// TIA Portal project "PalletizerLine" (V17)

(* hardware
DEVICE "S7-1500 station"  S7-1500 station
   slot 0: "Rail_0"  Rack  6ES7 590-1***0-0AA0
   slot 0: "PM 70W 120/230VAC"  PM 70W 120/230VAC  6EP1332-4BA00
   slot 1: "PLC_1"  CPU 1511-1 PN  6ES7 511-1AK02-0AB0  V2.9
      slot 3: "CPU display_1"  6ES7591-1AA00-0AA0
      slot 32768: "PROFINET interface_1"  X1
      slot 34817: "Virtual CP interface port_1"  Virtual CP interface port  Virtual CP interface port
   slot 2: "AI 8xU/I/RTD/TC ST_1"  AI 8xU/I/RTD/TC ST  6ES7 531-7KF00-0AB0  V2.2
   slot 3: "AI 8xU/I/RTD/TC ST_2"  AI 8xU/I/RTD/TC ST  6ES7 531-7KF00-0AB0  V2.2
   slot 4: "AI 8xU/I/RTD/TC ST_3"  AI 8xU/I/RTD/TC ST  6ES7 531-7KF00-0AB0  V2.2
   slot 5: "AI 8xU/I/RTD/TC ST_4"  AI 8xU/I/RTD/TC ST  6ES7 531-7KF00-0AB0  V2.2
   slot 6: "DI 16x24VDC BA_1"  DI 16x24VDC BA  6ES7 521-1BH10-0AA0  V1.1
DEVICE "HMI_TP1200"  TP1200 Comfort
   slot 0: "TP1200 Comfort"  TP1200 Comfort  6AV2 124-0MC01-0AX0  14.0.1.0
   slot 1: "HMI_RT_1"  TP1200 Comfort  6AV2 124-0MC01-0AX0  14.0.1.0
   slot 5: "Labeler HMI_TP1200.HMI.1"  PROFINET Interface  IE_CP  14.0.1.0
      slot 1: "PROFINET_Interface_1"  PROFINET Interface
         slot 1: "PORT_1"  Port  1.0.0.0
         slot 2: "PORT_2"  Port  1.0.0.0
   slot 7: "Labeler HMI_TP1200.HMI._CP_1"  MPI/DP Interface  MPI-DP_CP  14.0.1.0
*)

// ===== PLC "PLC_1"  CPU 1511-1 PN =====

VAR_GLOBAL   // PLC tag table "Default tag table"
   "System_Byte" AT %MB0 : Byte;   // System byte
   "FirstScan" AT %M0.0 : Bool;   // First scan PLC
   "DiagStatusUpdate" AT %M0.1 : Bool;   // Diagnostic status PLC updated
   "AlwaysTRUE" AT %M0.2 : Bool;   // Bit always true
   "AlwaysFALSE" AT %M0.3 : Bool;   // Bit always false
   "Clock_Byte" AT %MB1 : Byte;   // Clock byte
   "Clock_10Hz" AT %M1.0 : Bool;   // Clock pulse period 0,1s
   "Clock_5Hz" AT %M1.1 : Bool;   // Clock pulse period 0,2s
   "Clock_2.5Hz" AT %M1.2 : Bool;   // Clock pulse period 0,4s
   "Clock_2Hz" AT %M1.3 : Bool;   // Clock pulse period 0,5s
   "Clock_1.25Hz" AT %M1.4 : Bool;   // Clock pulse period 0,8s
   "Clock_1Hz" AT %M1.5 : Bool;   // Clock pulse period 1s
   "Clock_0.625Hz" AT %M1.6 : Bool;   // Clock pulse period 1,6s
   "Clock_0.5Hz" AT %M1.7 : Bool;   // Clock pulse period 2s
   "Tag_1" AT %I0.0 : Bool;
   "Tag_2" AT %Q0.0 : Bool;
   "Tag_3" AT %I0.1 : Bool;
   "Tag_4" AT %Q0.1 : Bool;
   "Tag_5" AT %Q0.2 : Bool;
   "Tag_6" AT %Q0.3 : Bool;
   "Tag_7" AT %Q0.4 : Bool;
   "Tag_8" AT %I0.2 : Bool;
   "Tag_9" AT %Q0.5 : Bool;
   "Tag_10" AT %I0.3 : Bool;
   "Tag_11" AT %Q0.6 : Bool;
   "Tag_12" AT %I0.4 : Bool;
   "Tag_13" AT %I0.5 : Bool;
   "Tag_14" AT %I0.6 : Bool;
   "Tag_15" AT %I0.7 : Bool;
   "Tag_16" AT %I1.0 : Bool;
   "Tag_17" AT %I1.1 : Bool;
   "Tag_18" AT %I1.2 : Bool;
   "Tag_19" AT %Q0.7 : Bool;
   "Tag_20" AT %Q1.0 : Bool;
   "Tag_21" AT %Q1.1 : Bool;
   "Tag_22" AT %Q1.2 : Bool;
   "Tag_23" AT %Q1.3 : Bool;
   "Tag_24" AT %Q1.4 : Bool;
   "Tag_25" AT %Q1.5 : Bool;
   "Tag_26" AT %Q1.6 : Bool;
   "Tag_27" AT %Q1.7 : Bool;
   "Tag_28" AT %Q2.0 : Bool;
   "Tag_29" AT %Q2.1 : Bool;
   "Tag_30" AT %Q2.2 : Bool;
   "Tag_31" AT %Q2.3 : Bool;
END_VAR

VAR_GLOBAL CONSTANT   // PLC tag table "CPG_Constants"
   "CPG_NO_OF_ELEMENTS_EVENT_STATUS_UPPER_LIM" : Int := 29;   // Number of Alarms, Warning and PackML Status events used by Event Status UDT (Array size of 0..x)
   "CPG_NO_OF_ADMIN_EVENTS_UPPER_LIM" : Int := 9;   // Number of Alarms and Warning events found in the PackTags Admin Area - active alarms / warnings. (Array size of 0..x)
   "CPG_NO_OF_ADMIN_EVENTS_HISTORY_UPPER_LIM" : Int := 9;   // Number of Alarms and Warning events found in the PackTags Admin Area - historical alarms / warnings. (Array size of 0..x)
   "CPG_NO_OF_PROD_CONSUMED_COUNT_UPPER_LIM" : Int := 0;   // Number of Prod Consumed Counter Array Size (PackTags Admin) (Array size of 0..x)
   "CPG_NO_OF_PROD_PROCESSED_COUNT_UPPER_LIM" : Int := 0;   // Number of Prod Processed Counter Array Size (PackTags Admin) (Array size of 0..x)
   "CPG_NO_OF_PROD_DEFECTIVE_COUNT_UPPER_LIM" : Int := 0;   // Number of Prod Defective Counter Array Size (PackTags Admin) (Array size of 0..x)
   "CPG_NO_OF_STS_ELEMENTS_EVENT_SUM_UPPER_LIM" : Int := 99;   // Number of Alarms, Warning and PackML Status events used by Event Summation UDT (Array size of 0..x)
   "CPG_NO_OF_HMI_SORT_EVENTS_UPPER_LIM" : Int := 19;   // Number of Alarms and Warning events found for the HMI area - sorted HMI alarms / warnings. (Array size of 0..x)
   "CPG_NO_OF_CFG_ALARMS_UPPER_LIM" : Int := 39;   // Number of Cfg Alarm event configurations (Array size of 0..x)
   "CPG_NO_OF_CFG_WARNINGS_UPPER_LIM" : Int := 29;   // Number of Cfg Warning event configurations (Array size of 0..x)
   "CPG_NO_OF_CFG_STATUS_UPPER_LIM" : Int := 19;   // Number of Cfg Status event configurations (Array size of 0..x)
   "CPG_NO_OF_STATUS_PARAMETERS_UPPER_LIM" : Int := 0;   // Number of Status Parameters (Array size of 0..x)
   "CPG_NO_OF_COMMAND_PARAMETERS_UPPER_LIM" : Int := 0;   // Number of Command Parameters (Array size of 0..x)
   "CPG_NO_OF_ADMIN_PARAMETERS_UPPER_LIM" : Int := 0;   // Number of Admin Parameters (Array size of 0..x)
   "CPG_NO_OF_RECIPE_UPPER_LIM" : Int := 20;   // Number of Project Recipies (Array size of 0..x)
   "CPG_NO_OF_SETPOINT_REAL_UPPER_LIM" : Int := 0;   // Number of Setpoints with a REAL type (Array size of 0..x)
   "CPG_NO_OF_SETPOINT_DINT_UPPER_LIM" : Int := 0;   // Number of Setpoints with a DINT type (Array size of 0..x)
   "CPG_NO_OF_SETPOINT_BOOL_UPPER_LIM" : Int := 0;   // Number of Setpoints with a BOOL type (Array size of 0..x)
   "CPG_NO_OF_SETPOINT_STRING_UPPER_LIM" : Int := 0;   // Number of Setpoints with a STRING type (Array size of 0..x)
   "CPG_PARTEO_NO_OF_ERRORS_UPPER_LIM" : Int := 100;   // Number of Unique Error IDs tracked by PARETO Error Blocks
END_VAR

VAR_GLOBAL CONSTANT   // PLC tag table "LPMLV30_Constants"
   "LPMLV30_MODE_INVALID" : DInt := 0;   // OMAC PackMLV30 unit mode Invalid
   "LPMLV30_MODE_PRODUCTION" : DInt := 1;   // OMAC PackMLV30 unit mode Production
   "LPMLV30_MODE_MAINTENANCE" : DInt := 2;   // OMAC PackMLV30 unit mode Maintenance
   "LPMLV30_MODE_MANUAL" : DInt := 3;   // OMAC PackMLV30 unit mode Manual
   "LPMLV30_MODE_USER_01" : DInt := 4;   // OMAC PackMLV30 user-defined unit mode 01
   "LPMLV30_MODE_USER_02" : DInt := 5;   // OMAC PackMLV30 user-defined unit mode 02
   "LPMLV30_MODE_USER_03" : DInt := 6;   // OMAC PackMLV30 user-defined unit mode 03
   "LPMLV30_MODE_USER_04" : DInt := 7;   // OMAC PackMLV30 user-defined unit mode 04
   "LPMLV30_MODE_USER_05" : DInt := 8;   // OMAC PackMLV30 user-defined unit mode 05
   "LPMLV30_MODE_USER_06" : DInt := 9;   // OMAC PackMLV30 user-defined unit mode 06
   "LPMLV30_MODE_USER_07" : DInt := 10;   // OMAC PackMLV30 user-defined unit mode 07
   "LPMLV30_MODE_USER_08" : DInt := 11;   // OMAC PackMLV30 user-defined unit mode 08
   "LPMLV30_MODE_USER_09" : DInt := 12;   // OMAC PackMLV30 user-defined unit mode 09
   "LPMLV30_MODE_USER_10" : DInt := 13;   // OMAC PackMLV30 user-defined unit mode 10
   "LPMLV30_MODE_USER_11" : DInt := 14;   // OMAC PackMLV30 user-defined unit mode 11
   "LPMLV30_MODE_USER_12" : DInt := 15;   // OMAC PackMLV30 user-defined unit mode 12
   "LPMLV30_MODE_USER_13" : DInt := 16;   // OMAC PackMLV30 user-defined unit mode 13
   "LPMLV30_MODE_USER_14" : DInt := 17;   // OMAC PackMLV30 user-defined unit mode 14
   "LPMLV30_MODE_USER_15" : DInt := 18;   // OMAC PackMLV30 user-defined unit mode 15
   "LPMLV30_MODE_USER_16" : DInt := 19;   // OMAC PackMLV30 user-defined unit mode 16
   "LPMLV30_MODE_USER_17" : DInt := 20;   // OMAC PackMLV30 user-defined unit mode 17
   "LPMLV30_MODE_USER_18" : DInt := 21;   // OMAC PackMLV30 user-defined unit mode 18
   "LPMLV30_MODE_USER_19" : DInt := 22;   // OMAC PackMLV30 user-defined unit mode 19
   "LPMLV30_MODE_USER_20" : DInt := 23;   // OMAC PackMLV30 user-defined unit mode 20
   "LPMLV30_MODE_USER_21" : DInt := 24;   // OMAC PackMLV30 user-defined unit mode 21
   "LPMLV30_MODE_USER_22" : DInt := 25;   // OMAC PackMLV30 user-defined unit mode 22
   "LPMLV30_MODE_USER_23" : DInt := 26;   // OMAC PackMLV30 user-defined unit mode 23
   "LPMLV30_MODE_USER_24" : DInt := 27;   // OMAC PackMLV30 user-defined unit mode 24
   "LPMLV30_MODE_USER_25" : DInt := 28;   // OMAC PackMLV30 user-defined unit mode 25
   "LPMLV30_MODE_USER_26" : DInt := 29;   // OMAC PackMLV30 user-defined unit mode 26
   "LPMLV30_MODE_USER_27" : DInt := 30;   // OMAC PackMLV30 user-defined unit mode 27
   "LPMLV30_MODE_USER_28" : DInt := 31;   // OMAC PackMLV30 user-defined unit mode 28
   "LPMLV30_STATE_UNDEFINED" : DInt := 0;   // OMAC PackMLV30 state Undefined
   "LPMLV30_STATE_CLEARING" : DInt := 1;   // OMAC PackMLV30 state Clearing
   "LPMLV30_STATE_STOPPED" : DInt := 2;   // OMAC PackMLV30 state Stopped
   "LPMLV30_STATE_STARTING" : DInt := 3;   // OMAC PackMLV30 state Starting
   "LPMLV30_STATE_IDLE" : DInt := 4;   // OMAC PackMLV30 state Idle
   "LPMLV30_STATE_SUSPENDED" : DInt := 5;   // OMAC PackMLV30 state Suspended
   "LPMLV30_STATE_EXECUTE" : DInt := 6;   // OMAC PackMLV30 state Execute
   "LPMLV30_STATE_STOPPING" : DInt := 7;   // OMAC PackMLV30 state Stopping
   "LPMLV30_STATE_ABORTING" : DInt := 8;   // OMAC PackMLV30 state Aborting
   "LPMLV30_STATE_ABORTED" : DInt := 9;   // OMAC PackMLV30 state Aborted
   "LPMLV30_STATE_HOLDING" : DInt := 10;   // OMAC PackMLV30 state Holding
   "LPMLV30_STATE_HELD" : DInt := 11;   // OMAC PackMLV30 state Held
   "LPMLV30_STATE_UNHOLDING" : DInt := 12;   // OMAC PackMLV30 state Unholding
   "LPMLV30_STATE_SUSPENDING" : DInt := 13;   // OMAC PackMLV30 state Suspending
   "LPMLV30_STATE_UNSUSPENDING" : DInt := 14;   // OMAC PackMLV30 state Unsuspending
   "LPMLV30_STATE_RESETTING" : DInt := 15;   // OMAC PackMLV30 state Resetting
   "LPMLV30_STATE_COMPLETING" : DInt := 16;   // OMAC PackMLV30 state Completing
   "LPMLV30_STATE_COMPLETE" : DInt := 17;   // OMAC PackMLV30 state Complete
   "LPMLV30_CMD_UNDEFINED" : DInt := 0;   // OMAC PackMLV30 control command Undefined
   "LPMLV30_CMD_RESET" : DInt := 1;   // OMAC PackMLV30 control command Reset
   "LPMLV30_CMD_START" : DInt := 2;   // OMAC PackMLV30 control command Start
   "LPMLV30_CMD_STOP" : DInt := 3;   // OMAC PackMLV30 control command Stop
   "LPMLV30_CMD_HOLD" : DInt := 4;   // OMAC PackMLV30 control command Hold
   "LPMLV30_CMD_UNHOLD" : DInt := 5;   // OMAC PackMLV30 control command Unhold
   "LPMLV30_CMD_SUSPEND" : DInt := 6;   // OMAC PackMLV30 control command Suspend
   "LPMLV30_CMD_UNSUSPEND" : DInt := 7;   // OMAC PackMLV30 control command Unsuspend
   "LPMLV30_CMD_ABORT" : DInt := 8;   // OMAC PackMLV30 control command Abort
   "LPMLV30_CMD_CLEAR" : DInt := 9;   // OMAC PackMLV30 control command Clear
   "LPMLV30_CMD_COMPLETE" : DInt := 10;   // OMAC PackMLV30 control command Complete
   "LPMLV30_LANGUAGE_1" : Int := 0;   // Texts in 1st language (default English)
   "LPMLV30_LANGUAGE_2" : Int := 1;   // Texts in 2nd language (default German)
   "LPMLV30_DIAG_BUFFER_UPPER_LIM" : Int := 15;   // Diagnostics buffer array upper boundary (0-based)
   "LPMLV30_LANGUAGES_UPPER_LIM" : Int := 2;   // (Number of languages - 1) -> Array[0..LPMLV30_LANGUAGES_UPPER_LIM]
   "LPMLV30_MODES_UPPER_LIM" : Int := 4;   // (Number of unit modes - 1) -> Array[0..LPMLV30_MODES_UPPER_LIM]
   "LPMLV30_STATES_UPPER_LIM" : Int := 17;   // (Number of states - 1) -> Array[0..LPMLV30_STATES_UPPER_LIM] (SHOULD ALWAYS BE 17!)
   "LPMLV30_MAX_MODES_UPPER_LIM" : Int := 31;   // (Maximum number of unit modes - 1) -> Array[0..LPMLV30_MAX_MODES_UPPER_LIM]
END_VAR

// folder: CPG_Types

TYPE "CPG_typePareto"
VERSION : 0.1
   STRUCT
      alarmID : DInt;
      alarmMessage : String[90];
      timesOccurred : UInt;   // number of times fault occurred
      totalDowntime : Real;   // total downtime resulting from all stops on this fault
      MTTR : Real;   // total downtime for this fault / total stops for this fault
      percentageOccurred : Real;   // total downtime on this fault / total downtime on whole machine
   END_STRUCT;
END_TYPE

TYPE "CPG_typeSortFilter"
   STRUCT
      cmdFilterActiveEvents : Bool;   // Filter for Active events: 1=only show active events; 0=show all events
      cmdFilterCategory : Bool;   // Filter by Category: filter events to show only selected category number
      cmdSortCategory : Bool;   // Sort by Category: 1=sort events by ascending category number
      cfgTimeSortDirection : Bool;   // Sort by Time: 1=newest first; 0=oldest first
      cfgEventListOffset : Int;   // Commanded event list offset (used for scrolling)
      cfgFilterCategory : Int;   // Filter by Category: filtered category number
   END_STRUCT;
END_TYPE

TYPE "CPG_typeRecipeSetpoint_BOOL"
   STRUCT
      IN : Bool;   // Incoming recipe value
      SaveSetpoint : Bool;   // Command to save current (out) value to current recipe
      RevertSetpoint : Bool;   // Command to revert current (out) value to saved value
      RecipeValues : Array[0.."CPG_NO_OF_RECIPE_UPPER_LIM"] of Bool;   // Saved value for all recipes
      SetpointName : Array[0.."LPMLV30_LANGUAGES_UPPER_LIM"] of String[60];   // Setpoint name in all languages
      Text_True : Array[0.."LPMLV30_LANGUAGES_UPPER_LIM"] of String[60];   // True text in all languages
      Text_False : Array[0.."LPMLV30_LANGUAGES_UPPER_LIM"] of String[60];   // False text in all languages
      CurrentName : String[60];   // Setpoint name for current language
      CurrentTextTrue : String[60];   // Text to display for a true value
      CurrentTextFalse : String[60];   // Text to display for a false value
      DisableRecipeControl : Bool;   // When true, the value is not treated like a recipe
      SetpointChangeEnabled : Bool;   // Changing the setpoint is possible
      SetpointChangeDisabled : Bool;   // Change not allowed because FB enable input is false
      RecipeSetpointDiff : Bool;   // Currently running (out) value not equal to saved recipe value
      OUT : Bool;   // Currently running, validated recipe value
      Out_Text : String[60];   // Display text for OUT
      CurrentRecipeValue : Bool;   // Current saved recipe value
      CurrentRecipeValue_Text : String[60];   // Display text for Current Recipe
      RecipeValueA : Bool;   // Value for recipe A
      RecipeA_Text : String[60];   // Display text for A
      RecipeValueB : Bool;   // Value for recipe B
      RecipeB_Text : String[60];   // Display text for B
      RecipeValueC : Bool;   // Value for recipe C
      RecipeC_Text : String[60];   // Display text for C
   END_STRUCT;
END_TYPE

TYPE "CPG_typeRecipeSetpoint_REAL"
   STRUCT
      IN : Real;   // Incoming recipe value
      SaveSetpoint : Bool;   // Command to save current (out) value to current recipe
      RevertSetpoint : Bool;   // Command to revert current (out) value to saved value
      RecipeValues : Array[0.."CPG_NO_OF_RECIPE_UPPER_LIM"] of Real;   // Saved value for all recipes
      SetpointName : Array[0.."LPMLV30_LANGUAGES_UPPER_LIM"] of String[60];   // Setpoint name in all languages
      CurrentName : String[60];   // Setpoint name for current language
      minLimit : Real;   // Minimum value for setpoint
      maxLimit : Real;   // Maximum value for setpoint
      unit : String[60];   // Units of measurement
      DisableRecipeControl : Bool;   // When true, the value is not treated like a recipe
      SetpointChangeEnabled : Bool;   // Changing the setpoint is possible
      SetpointChangeDisabled : Bool;   // Change not allowed because FB enable input is false
      RecipeSetpointDiff : Bool;   // Currently running (out) value not equal to saved recipe value
      minLimitReached : Bool;   // IN value was below minimum
      maxLimitReached : Bool;   // IN value was above maximum
      OUT : Real;   // Currently running, validated recipe value
      CurrentRecipeValue : Real;   // Current saved recipe value
      RecipeValueA : Real;   // Value for recipe A
      RecipeValueB : Real;   // Value for recipe B
      RecipeValueC : Real;   // Value for recipe C
   END_STRUCT;
END_TYPE

TYPE "CPG_typeRecipeSetpoint_DINT"
   STRUCT
      IN : DInt;   // Incoming recipe value
      SaveSetpoint : Bool;   // Command to save current (out) value to current recipe
      RevertSetpoint : Bool;   // Command to revert current (out) value to saved value
      RecipeValues : Array[0.."CPG_NO_OF_RECIPE_UPPER_LIM"] of DInt;   // Saved value for all recipes
      SetpointName : Array[0.."LPMLV30_LANGUAGES_UPPER_LIM"] of String[60];   // Setpoint name in all languages
      CurrentName : String[60];   // Setpoint name for current language
      minLimit : DInt;   // Minimum value for setpoint
      maxLimit : DInt;   // Maximum value for setpoint
      unit : String[60];   // Units of measurement
      DisableRecipeControl : Bool;   // When true, the value is not treated like a recipe
      SetpointChangeEnabled : Bool;   // Changing the setpoint is possible
      SetpointChangeDisabled : Bool;   // Change not allowed because FB enable input is false
      RecipeSetpointDiff : Bool;   // Currently running (out) value not equal to saved recipe value
      minLimitReached : Bool;   // IN value was below minimum
      maxLimitReached : Bool;   // IN value was above maximum
      OUT : DInt;   // Currently running, validated recipe value
      CurrentRecipeValue : DInt;   // Current saved recipe value
      RecipeValueA : DInt;   // Value for recipe A
      RecipeValueB : DInt;   // Value for recipe B
      RecipeValueC : DInt;   // Value for recipe C
   END_STRUCT;
END_TYPE

TYPE "CPG_typeRecipeSetpoint_STRING"
   STRUCT
      IN : String[60];   // Incoming recipe value
      SaveSetpoint : Bool;   // Command to save current (out) value to current recipe
      RevertSetpoint : Bool;   // Command to revert current (out) value to saved value
      RecipeValues : Array[0.."CPG_NO_OF_RECIPE_UPPER_LIM"] of String[60];   // Saved value for all recipes
      SetpointName : Array[0.."LPMLV30_LANGUAGES_UPPER_LIM"] of String[60];   // Setpoint name in all languages
      CurrentSetpointName : String[60];   // Setpoint name for current language
      DisableRecipeControl : Bool;   // When true, the value is not treated like a recipe
      SetpointChangeEnabled : Bool;   // Changing the setpoint is possible
      SetpointChangeDisabled : Bool;   // Change not allowed because FB enable input is false
      RecipeSetpointDiff : Bool;   // Currently running (out) value not equal to saved recipe value
      OUT : String[60];   // Currently running, validated recipe value
      CurrentRecipeValue : String[60];   // Current saved recipe value
      RecipeValueA : String[60];   // Value for recipe A
      RecipeValueB : String[60];   // Value for recipe B
      RecipeValueC : String[60];   // Value for recipe C
   END_STRUCT;
END_TYPE

TYPE "CPG_typeParameter(Real)"
VERSION : 0.1
   STRUCT
      ID : DInt;   // Parameter ID - This is the arbitrary (user defined) ID value of the parameter
      "Name" : String[24];   // Parameter Name - The literal parameter name is used to describe the parameter number and its associated value (e.g. Glue Temp)
      Unit : String[5];   // Parameter Unit of Measure - The parameter unit is used to describe the unit of measure of the parameter and its associated value (e.g. DegF)
      Value : Real;   // Parameter Value - This is the numeric or string value of the parameter (e.g. 100.2)
   END_STRUCT;
END_TYPE

TYPE "CPG_typeParameter(DINT)"
VERSION : 0.1
   STRUCT
      ID : DInt;   // Parameter ID - This is the arbitrary (user defined) ID value of the parameter
      "Name" : String[24];   // Parameter Name - The literal parameter name is used to describe the parameter number and its associated value (e.g. Glue Temp)
      Unit : String[5];   // Parameter Unit of Measure - The parameter unit is used to describe the unit of measure of the parameter and its associated value (e.g. DegF)
      Value : DInt;   // Parameter Value - This is the numeric or string value of the parameter (e.g. 100)
   END_STRUCT;
END_TYPE

TYPE "CPG_typeParameter(String)"
VERSION : 0.1
   STRUCT
      ID : DInt;   // Parameter ID - This is the arbitrary (user defined) ID value of the parameter
      "Name" : String[24];   // Parameter Name - The literal parameter name is used to describe the parameter number and its associated value (e.g. Glue Temp)
      Unit : String[5];   // Parameter Unit of Measure - The parameter unit is used to describe the unit of measure of the parameter and its associated value (e.g. DegF)
      Value : String[24];   // Parameter Value - This is the numeric or string value of the parameter (e.g. '6ES7518-4AP00-0AB0')
   END_STRUCT;
END_TYPE

TYPE "CPG_typeProdCount(DINT)"
VERSION : 0.1
   STRUCT
      ID : DInt;   // Product ID - This is the arbitrary (user defined) ID value of the consumed production material
      "Name" : String[24];   // Descriptive name - The name is used to literally describe the material ID, and its associated material
      Unit : String[5];   // Unit of measure - The unit tag is used to describe the names associated with a specific material used by the machine
      Count : DInt;   // Value - The count value is used as a variable for displaying information about the amount of consumed
      AccCount : DInt;   // Value - The accumulative count value is used as a variable for displaying information about the total amount of consumed production material
   END_STRUCT;
END_TYPE

TYPE "CPG_typeRecipeControl"
   STRUCT
      CurrentRecipeID : Int;   // The ID of the currently loaded recipe
      CurrentRecipeName : String[60];   // The name of the currently loaded recipe
      RecipeChange : Bool;   // Bit is true if a recipe change is in progress
      RecipeChangeNum : Int;   // Work variable, do not modify
      RecipeSave : Bool;   // Bit is true if a recipe save or saveas is in progress
      RecipeSaveNum : Int;   // Work variable, do not modify
      RecipeCopy : Bool;   // Bit is true if a recipe copy is in progress
      RecipeCopyNum : Int;   // Work variable, do not modify
      RecipeDelete : Bool;   // Bit is true if a recipe delete is in progress
      RecipeDeleteNum : Int;   // Work variable, do not modify
      RecipeSourceID : Int;   // In a copy or save, this is the ID of the recipe souce
      RecipeDestinationID : Int;   // In a copy, save, or delete, this is the ID of the recipe to be overwritten
      LanguageSelection : Int;   // The currently selected language
      RecipeSetpointDiff : Bool;   // At least one setpoint's value is different from the currently loaded recipe
      RecipeChangeDisabled : Bool;   // Bit is true if "Enable" input to Recipe Control FB is false
      RecipeID_A : Int;   // ID of recipe A
      RecipeName_A : String[60];   // Name of recipe A
      RecipeID_B : Int;   // ID of recipe B
      RecipeName_B : String[60];   // Name of recipe B
      RecipeID_C : Int;   // ID of recipe C
      RecipeName_C : String[60];   // Name of recipe C
   END_STRUCT;
END_TYPE

TYPE "CPG_typeEventStatus"
AUTHOR : FoodBev
FAMILY : ISATR88e
NAME : EventSts
VERSION : 1.0
   STRUCT
      sts_FirstOutEvent : "CPG_typeEvent";   // Event Info of the very first active event (irregardeless of the cat)
      sts_FirstOutEventCat : Array[0..9] of "CPG_typeEvent";
      sts_Events : Array[0.."CPG_NO_OF_ELEMENTS_EVENT_STATUS_UPPER_LIM"] of "CPG_typeEvent";
      sts_NumEvents : Int;   // Number of all current active events
      sts_NumAllEvents : Int;   // Number of all current events
      out_ZeroEvent : "CPG_typeEvent";   // null event information
      sts_Category_0_Latched : Bool;   // Category 0 Event - latched (require reset cmd)
      sts_Category_1_Latched : Bool;   // Category 1 Event - latched (require reset cmd)
      sts_Category_2_Latched : Bool;   // Category 2 Event - latched (require reset cmd)
      sts_Category_3_Latched : Bool;   // Category 3 Event - latched (require reset cmd)
      sts_Category_4_Latched : Bool;   // Category 4 Event - latched (require reset cmd)
      sts_Category_5_Latched : Bool;   // Category 5 Event - latched (require reset cmd)
      sts_Category_6_Latched : Bool;   // Category 6 Event - latched (require reset cmd)
      sts_Category_7_Latched : Bool;   // Category 7 Event - latched (require reset cmd)
      sts_Category_8_Latched : Bool;   // Category 8 Event - latched (require reset cmd)
      sts_Category_9_Latched : Bool;   // Category 9 Event - latched (require reset cmd)
      sts_Category_0_NotLatched : Bool;   // Category 0 Event - NotLatched (currently active)
      sts_Category_1_NotLatched : Bool;   // Category 1 Event - NotLatched (currently active)
      sts_Category_2_NotLatched : Bool;   // Category 2 Event - NotLatched (currently active)
      sts_Category_3_NotLatched : Bool;   // Category 3 Event - NotLatched (currently active)
      sts_Category_4_NotLatched : Bool;   // Category 4 Event - NotLatched (currently active)
      sts_Category_5_NotLatched : Bool;   // Category 5 Event - NotLatched (currently active)
      sts_Category_6_NotLatched : Bool;   // Category 6 Event - NotLatched (currently active)
      sts_Category_7_NotLatched : Bool;   // Category 7 Event - NotLatched (currently active)
      sts_Category_8_NotLatched : Bool;   // Category 8 Event - NotLatched (currently active)
      sts_Category_9_NotLatched : Bool;   // Category 9 Event - NotLatched (currently active)
      sts_CurrentActiveEvent : Bool;   // Active # of Event
      wrk_ResetID : Int;   // Working Variable - DO NOT MODIFY
      wrk_EventArraySize : Int;   // Working Variable - DO NOT MODIFY
      wrk_UpdateEventListID : Int;   // Working Variable - DO NOT MODIFY
      wrk_LanguageSelection : Int;   // This is the value of language selected in the HMI
      wrk_MessagePrefix : String[10];   // Working Variable - DO NOT MODIFY
   END_STRUCT;
END_TYPE

TYPE "CPG_typeEventCfg"
AUTHOR : FoodBev
FAMILY : ISATR88e
NAME : EvntCfgA
VERSION : 1.0
   STRUCT
      ID : Int;   // ID Value - from PackTags Reason Code, 1=E-Stop pushed, 3=Main off, etc.
      value : Int;   // Reason Code 'Value' - allows for detailed breakdown of ID, ie 1=Discharge,
      message : Array[0.."LPMLV30_LANGUAGES_UPPER_LIM"] of String[60];   // Alarm Message - 0=English, 1=German, 2=Spanish, 3=Italian, 4=French
      category : Int;   // Category Value (0-9)
   END_STRUCT;
END_TYPE

TYPE "CPG_typeEvent"
AUTHOR : FoodBev
FAMILY : ISATR88e
NAME : Event
VERSION : 1.0
   STRUCT
      Trigger : Bool;   // 1=Alarm is currently active
      ID : DInt;   // Alarm Message Identification Number, see PackTags Reason Code (e.g. 1=E-Stop pushed, 3=Mains turned off, etc.)
      Value : DInt;   // Alarm Mesage Value to break down the Alarm.ID to greater detail
      Message : String[60];   // Alarm Message Text (= message prefix + alarm message)
      Category : DInt;   // Alarm Category Value (0-9)
      DateTime : Array[0..6] of DInt;   // Date and Time the Event Occurred
      DateTimeDTL : DTL;   // Date and LTime (DTL) the event was initially triggered (date and time-of-day information in nanoseconds since 01/01/1970 0:0)
      AckDateTime : Array[0..6] of DInt;   // Date and Time the Event was Acknowledged
      AckDateTimeDTL : DTL;   // Date and LTime (DTL) the event was acknowledged (date and time-of-day information in nanoseconds since 01/01/1970 0:0)
   END_STRUCT;
   // // DateTime[0] : Year
   // // DateTime[1] : Month
   // // DateTime[2] : Day
   // // DateTime[3] : Hour (24hr format)
   // // DateTime[4] : Min
   // // DateTime[5] : Sec
   // // DateTime[6] : USec (1/1,000,000 sec)
   // // AckDateTime[0] : Year
   // // AckDateTime[1] : Month
   // // AckDateTime[2] : Day
   // // AckDateTime[3] : Hour (24hr format)
   // // AckDateTime[4] : Min
   // // AckDateTime[5] : Sec
   // // AckDateTime[6] : USec (1/1,000,000 sec)
END_TYPE

TYPE "CPG_typeEventSummation"
AUTHOR : FoodBev
FAMILY : ISATR88e
NAME : EventSum
VERSION : 1.0
   STRUCT
      sts_FirstOutEvent : "CPG_typeEvent";   // First Out (Stop Reason) Event
      sts_FirstOutEventCat : Array[0..9] of "CPG_typeEvent";   // First Out (Stop Reason) Event by Category\
      sts_Events : Array[0.."CPG_NO_OF_STS_ELEMENTS_EVENT_SUM_UPPER_LIM"] of "CPG_typeEvent";   // All Active Events
      sts_NumEvents : Int;   // Number of Active Events
      sts_Category_0_Latched : Bool;   // Category 0 Event - latched (require reset cmd)
      sts_Category_1_Latched : Bool;   // Category 1 Event - latched (require reset cmd)
      sts_Category_2_Latched : Bool;   // Category 2 Event - latched (require reset cmd)
      sts_Category_3_Latched : Bool;   // Category 3 Event - latched (require reset cmd)
      sts_Category_4_Latched : Bool;   // Category 4 Event - latched (require reset cmd)
      sts_Category_5_Latched : Bool;   // Category 5 Event - latched (require reset cmd)
      sts_Category_6_Latched : Bool;   // Category 6 Event - latched (require reset cmd)
      sts_Category_7_Latched : Bool;   // Category 7 Event - latched (require reset cmd)
      sts_Category_8_Latched : Bool;   // Category 8 Event - latched (require reset cmd)
      sts_Category_9_Latched : Bool;   // Category 9 Event - latched (require reset cmd)
      sts_Category_0_NotLatched : Bool;   // Category 0 Event - NotLatched (currently active)
      sts_Category_1_NotLatched : Bool;   // Category 1 Event - NotLatched (currently active)
      sts_Category_2_NotLatched : Bool;   // Category 2 Event - NotLatched (currently active)
      sts_Category_3_NotLatched : Bool;   // Category 3 Event - NotLatched (currently active)
      sts_Category_4_NotLatched : Bool;   // Category 4 Event - NotLatched (currently active)
      sts_Category_5_NotLatched : Bool;   // Category 5 Event - NotLatched (currently active)
      sts_Category_6_NotLatched : Bool;   // Category 6 Event - NotLatched (currently active)
      sts_Category_7_NotLatched : Bool;   // Category 7 Event - NotLatched (currently active)
      sts_Category_8_NotLatched : Bool;   // Category 8 Event - NotLatched (currently active)
      sts_Category_9_NotLatched : Bool;   // Category 9 Event - NotLatched (currently active)
      sts_CurrentActiveEvent : Bool;   // Event Active = 1, not active = 0
      wrk_EventArraySize : Int;   // Maximum Array Size - DO NOT MODIFY
      wrk_Category_0_Latched : Bool;   // Working Variable - DO NOT MODIFY
      wrk_Category_1_Latched : Bool;   // Working Variable - DO NOT MODIFY
      wrk_Category_2_Latched : Bool;   // Working Variable - DO NOT MODIFY
      wrk_Category_3_Latched : Bool;   // Working Variable - DO NOT MODIFY
      wrk_Category_4_Latched : Bool;   // Working Variable - DO NOT MODIFY
      wrk_Category_5_Latched : Bool;   // Working Variable - DO NOT MODIFY
      wrk_Category_6_Latched : Bool;   // Working Variable - DO NOT MODIFY
      wrk_Category_7_Latched : Bool;   // Working Variable - DO NOT MODIFY
      wrk_Category_8_Latched : Bool;   // Working Variable - DO NOT MODIFY
      wrk_Category_9_Latched : Bool;   // Working Variable - DO NOT MODIFY
      wrk_Category_0_NotLatched : Bool;   // Working Variable - DO NOT MODIFY
      wrk_Category_1_NotLatched : Bool;   // Working Variable - DO NOT MODIFY
      wrk_Category_2_NotLatched : Bool;   // Working Variable - DO NOT MODIFY
      wrk_Category_3_NotLatched : Bool;   // Working Variable - DO NOT MODIFY
      wrk_Category_4_NotLatched : Bool;   // Working Variable - DO NOT MODIFY
      wrk_Category_5_NotLatched : Bool;   // Working Variable - DO NOT MODIFY
      wrk_Category_6_NotLatched : Bool;   // Working Variable - DO NOT MODIFY
      wrk_Category_7_NotLatched : Bool;   // Working Variable - DO NOT MODIFY
      wrk_Category_8_NotLatched : Bool;   // Working Variable - DO NOT MODIFY
      wrk_Category_9_NotLatched : Bool;   // Working Variable - DO NOT MODIFY
      wrk_CurrentActiveEvent : Bool;   // Working Variable - DO NOT MODIFY
   END_STRUCT;
END_TYPE

TYPE "CPG_typePackML_ModuleSts"
AUTHOR : FoodBev
FAMILY : ISATR88e
NAME : PML_MdSt
VERSION : 1.0
   STRUCT
      cmd_Reset : Bool;   // Reset
      sts_Resetting_SC : Bool;   // Resetting State Complete
      cmd_Start : Bool;   // Start
      sts_Starting_SC : Bool;   // Starting State Complete
      cmd_Stop : Bool;   // Stop
      sts_Stopping_SC : Bool;   // Stopping State Complete
      cmd_Hold : Bool;   // Hold
      sts_Holding_SC : Bool;   // Holding State Complete
      cmd_UnHold : Bool;   // UnHold
      sts_UnHolding_SC : Bool;   // UnHolding State Complete
      cmd_Suspend : Bool;   // Suspend
      sts_Suspending_SC : Bool;   // Suspending State Complete
      cmd_UnSuspend : Bool;   // UnSuspend
      sts_UnSuspending_SC : Bool;   // UnSuspending State Complete
      cmd_Abort : Bool;   // Abort
      sts_Aborting_SC : Bool;   // Aborting State Complete
      cmd_Clear : Bool;   // Clear
      sts_Clearing_SC : Bool;   // Clearing State Complete
      sts_Execute_SC : Bool;   // Execute State Complete
      sts_Completing_SC : Bool;   // Completing State Complete
      moduleActive : Bool;   // Module Active Bit
      ONS : Bool;   // Internal One Shot Bit - Do not modify
   END_STRUCT;
END_TYPE

TYPE "CPG_typeMessagePrefix"
VERSION : 0.1
   STRUCT
      messagePrefix : Array[0.."LPMLV30_LANGUAGES_UPPER_LIM"] of String[30];   // Multi-Lingual Message for Prefix (i.e 0=EN, 1=DE, 2=SP/ES, 3=IT, 4=FR)
   END_STRUCT;
END_TYPE

// folder: LPMLV30_Types

TYPE "typeLPMLV30_DiagnosticsEntry"
TITLE = typeLPMLV30_DiagnosticsEntry
VERSION : 0.1
// Support: tech.team.motioncontrol@siemens.com 
// Fax: +49 (0) 9131/98-1297
   STRUCT
      timestamp : DTL := DTL#1970-01-01-00:00:00;   // Timestamp for this entry
      UnitModeCurrent : Byte := 16#00;   // Current unit mode
      StateCurrent : Byte := 16#00;   // Current state
      UnitMode : Byte := 16#00;   // Requested unit mode
      CntrlCmd : Byte := 16#00;   // Request control command
      SC : Bool := false;   // State complete signal
      message : Byte := 16#00;   // Message for this entry
   END_STRUCT;
END_TYPE

TYPE "typeLPMLV30_Configuration"
TITLE = typeLPMLV30_Configuration
VERSION : 0.1
// Support: tech.team.motioncontrol@siemens.com 
// Fax: +49 (0) 9131/98-1297
   STRUCT
      disabledUnitModes : Array[0.."LPMLV30_MAX_MODES_UPPER_LIM"] of Bool;   // TRUE: Disable unit mode xx
      disabledStatesInUnitModes : Array[0.."LPMLV30_MAX_MODES_UPPER_LIM"] of DInt;   // TRUE: Disable states in unit mode (bit number = state number)
   END_STRUCT;
   // disabledUnitModes[4] := false;
   // disabledUnitModes[5] := false;
   // disabledUnitModes[6] := false;
   // disabledUnitModes[7] := false;
   // disabledUnitModes[8] := false;
   // disabledUnitModes[0] := false;
   // disabledUnitModes[1] := false;
   // disabledUnitModes[2] := false;
   // disabledUnitModes[3] := false;
   // disabledUnitModes[9] := false;
   // disabledUnitModes[10] := false;
   // disabledUnitModes[11] := false;
   // disabledUnitModes[12] := true;
   // disabledUnitModes[13] := true;
   // disabledUnitModes[14] := true;
   // disabledUnitModes[15] := true;
   // disabledUnitModes[16] := true;
   // disabledUnitModes[17] := true;
   // disabledUnitModes[18] := true;
   // disabledUnitModes[19] := true;
   // disabledUnitModes[20] := true;
   // disabledUnitModes[21] := true;
   // disabledUnitModes[22] := true;
   // disabledUnitModes[23] := true;
   // disabledUnitModes[24] := true;
   // disabledUnitModes[25] := true;
   // disabledUnitModes[26] := true;
   // disabledUnitModes[27] := true;
   // disabledUnitModes[28] := true;
   // disabledUnitModes[29] := true;
   // disabledUnitModes[30] := true;
   // disabledUnitModes[31] := true;
   // disabledStatesInUnitModes[0] := 0;
   // disabledStatesInUnitModes[1] := 0;
   // disabledStatesInUnitModes[2] := 0;
   // disabledStatesInUnitModes[3] := 0;
   // disabledStatesInUnitModes[4] := 0;
   // disabledStatesInUnitModes[5] := 0;
   // disabledStatesInUnitModes[6] := 0;
   // disabledStatesInUnitModes[7] := 0;
   // disabledStatesInUnitModes[8] := 0;
   // disabledStatesInUnitModes[9] := 0;
   // disabledStatesInUnitModes[10] := 0;
   // disabledStatesInUnitModes[11] := 0;
   // disabledStatesInUnitModes[12] := 0;
   // disabledStatesInUnitModes[13] := 0;
   // disabledStatesInUnitModes[14] := 0;
   // disabledStatesInUnitModes[15] := 0;
   // disabledStatesInUnitModes[16] := 0;
   // disabledStatesInUnitModes[17] := 0;
   // disabledStatesInUnitModes[18] := 0;
   // disabledStatesInUnitModes[19] := 0;
   // disabledStatesInUnitModes[20] := 0;
   // disabledStatesInUnitModes[21] := 0;
   // disabledStatesInUnitModes[22] := 0;
   // disabledStatesInUnitModes[23] := 0;
   // disabledStatesInUnitModes[24] := 0;
   // disabledStatesInUnitModes[25] := 0;
   // disabledStatesInUnitModes[26] := 0;
   // disabledStatesInUnitModes[27] := 0;
   // disabledStatesInUnitModes[28] := 0;
   // disabledStatesInUnitModes[29] := 0;
   // disabledStatesInUnitModes[30] := 0;
   // disabledStatesInUnitModes[31] := 0;
END_TYPE

TYPE "typeLPMLV30_Diagnostics"
TITLE = typeLPMLV30_Diagnostics
VERSION : 0.1
// Support: tech.team.motioncontrol@siemens.com 
// Fax: +49 (0) 9131/98-1297
   STRUCT
      bufferIndex : Int := -1;   // Index of actual buffer entry
      buffer : Array[0.."LPMLV30_DIAG_BUFFER_UPPER_LIM"] of "typeLPMLV30_DiagnosticsEntry";   // Diagnostics information buffer
   END_STRUCT;
END_TYPE

TYPE "typeLPMLV30_NamesConfiguration"
TITLE = typeLPMLV30_NamesConfiguration
VERSION : 0.1
// Support: tech.team.motioncontrol@siemens.com 
// Fax: +49 (0) 9131/98-1297
   STRUCT
      unitModesNames : Array[0.."LPMLV30_LANGUAGES_UPPER_LIM", 0.."LPMLV30_MODES_UPPER_LIM"] of String[18];   // Names of unit modes [First index language, Second unit mode no]
      statesNames : Array[0.."LPMLV30_LANGUAGES_UPPER_LIM", 0.."LPMLV30_STATES_UPPER_LIM"] of String[16];   // Names of states [First index language, Second state no]
   END_STRUCT;
   // statesNames[0,0] := 'Undefined';
   // statesNames[0,1] := 'Clearing';
   // statesNames[0,2] := 'Stopped';
   // statesNames[0,3] := 'Starting';
   // statesNames[0,4] := 'Idle';
   // statesNames[0,5] := 'Suspended';
   // statesNames[0,6] := 'Execute';
   // statesNames[0,7] := 'Stopping';
   // statesNames[0,8] := 'Aborting';
   // statesNames[0,9] := 'Aborted';
   // statesNames[0,10] := 'Holding';
   // statesNames[0,11] := 'Held';
   // statesNames[0,12] := 'UnHolding';
   // statesNames[0,13] := 'Suspending';
   // statesNames[0,14] := 'UnSuspending';
   // statesNames[0,15] := 'Resetting';
   // statesNames[0,16] := 'Completing';
   // statesNames[0,17] := 'Complete';
   // statesNames[1,0] := 'Undefiniert';
   // statesNames[1,1] := 'Clearing';
   // statesNames[1,2] := 'Stopped';
   // statesNames[1,3] := 'Starting';
   // statesNames[1,4] := 'Idle';
   // statesNames[1,5] := 'Suspended';
   // statesNames[1,6] := 'Execute';
   // statesNames[1,7] := 'Stopping';
   // statesNames[1,8] := 'Aborting';
   // statesNames[1,9] := 'Aborted';
   // statesNames[1,10] := 'Holding';
   // statesNames[1,11] := 'Held';
   // statesNames[1,12] := 'UnHolding';
   // statesNames[1,13] := 'Suspending';
   // statesNames[1,14] := 'UnSuspending';
   // statesNames[1,15] := 'Resetting';
   // statesNames[1,16] := 'Completing';
   // statesNames[1,17] := 'Complete';
   // unitModesNames[0,0] := 'Invalid';
   // unitModesNames[0,1] := 'Production';
   // unitModesNames[0,2] := 'Maintenance';
   // unitModesNames[0,3] := 'Manual';
   // unitModesNames[0,4] := 'User Mode 01';
   // unitModesNames[1,0] := 'Undefiniert';
   // unitModesNames[1,1] := 'Produktion';
   // unitModesNames[1,2] := 'Wartung';
   // unitModesNames[1,3] := 'Hand';
   // unitModesNames[1,4] := 'Benutzer Mode 01';
END_TYPE

// folder: EM00_Transport

DATA_BLOCK "EM00"   // DB31649
TITLE = EM00
{ S7_Optimized_Access := 'TRUE' }
AUTHOR : tech.team.motioncontrol@siemens.com
FAMILY : CPG
VERSION : 1.1
// Support: tech.team.motioncontrol@siemens.com
   VAR
      PackML_Sts : Struct   // PackML Module Status - EM and all control modules
         Unit : "CPG_typePackML_ModuleSts";   // PackML Module Status - EM - master status
         Alarm : "CPG_typePackML_ModuleSts";   // PackML Module Status - alarm status
         CM01 : "CPG_typePackML_ModuleSts";   // PackML Module Status - CM 01
         CM02 : "CPG_typePackML_ModuleSts";   // PackML Module Status - CM 02
         CM03 : "CPG_typePackML_ModuleSts";   // PackML Module Status - CM 03
         CM04 : "CPG_typePackML_ModuleSts";   // PackML Module Status - CM 04
         CM05 : "CPG_typePackML_ModuleSts";   // PackML Module Status - CM 05
         CM06 : "CPG_typePackML_ModuleSts";   // PackML Module Status - CM 06
         CM07 : "CPG_typePackML_ModuleSts";   // PackML Module Status - CM 07
         CM08 : "CPG_typePackML_ModuleSts";   // PackML Module Status - CM 08
         CM09 : "CPG_typePackML_ModuleSts";   // PackML Module Status - CM 09
         CM10 : "CPG_typePackML_ModuleSts";   // PackML Module Status - CM 10
      END_STRUCT;
      Alarm : "CPG_typeEventStatus";   // Alarm Event Status - EM00 Status
      Warning : "CPG_typeEventStatus";   // Warning Event Status - EM00 Status
      Status : "CPG_typeEventStatus";   // Event Status - EM00 Status
   END_VAR
BEGIN
END_DATA_BLOCK

// folder: EM00_Transport/Instances

DATA_BLOCK "InstEM00_00_Main"   // DB31640
TITLE = instEM00_00_Main
{ S7_Optimized_Access := 'TRUE' }
AUTHOR : tech.team.motioncontrol@siemens.com
FAMILY : CPG
VERSION : 1.0
// Support: tech.team.motioncontrol@siemens.com
// Fax: +49 (0) 9131/98-1297
// stored: InstanceOfName EM00_00_Main
"EM00_00_Main"
BEGIN
END_DATA_BLOCK

// folder: EM01_Palletizing

DATA_BLOCK "EM01"   // DB31669
TITLE = EM01
{ S7_Optimized_Access := 'TRUE' }
AUTHOR : tech.team.motioncontrol@siemens.com
FAMILY : CPG
VERSION : 1.0
// Support: tech.team.motioncontrol@siemens.com
// Fax: +49 (0) 9131/98-1297
   VAR
      PackML_Sts : Struct   // PackML Module Status - EM and all control modules
         Unit : "CPG_typePackML_ModuleSts";   // PackML Module Status - EM - master status
         Alarm : "CPG_typePackML_ModuleSts";   // PackML Module Status - alarm status
         CM01 : "CPG_typePackML_ModuleSts";   // PackML Module Status - CM 01
         CM02 : "CPG_typePackML_ModuleSts";   // PackML Module Status - CM 02
         CM03 : "CPG_typePackML_ModuleSts";   // PackML Module Status - CM 03
         CM04 : "CPG_typePackML_ModuleSts";   // PackML Module Status - CM 04
         CM05 : "CPG_typePackML_ModuleSts";   // PackML Module Status - CM 05
         CM06 : "CPG_typePackML_ModuleSts";   // PackML Module Status - CM 06
         CM07 : "CPG_typePackML_ModuleSts";   // PackML Module Status - CM 07
         CM08 : "CPG_typePackML_ModuleSts";   // PackML Module Status - CM 08
         CM09 : "CPG_typePackML_ModuleSts";   // PackML Module Status - CM 09
         CM10 : "CPG_typePackML_ModuleSts";   // PackML Module Status - CM 10
      END_STRUCT;
      Alarm : "CPG_typeEventStatus";   // Alarm Event Status - EM01 Status
      Warning : "CPG_typeEventStatus";   // Warning Event Status - EM01 Status
      Status : "CPG_typeEventStatus";   // Event Status - EM01 Status
   END_VAR
BEGIN
END_DATA_BLOCK

// folder: EM01_Palletizing/Instances

DATA_BLOCK "InstEM01_00_Main"   // DB31660
TITLE = InstEM01_00_Main
{ S7_Optimized_Access := 'TRUE' }
AUTHOR : tech.team.motioncontrol@siemens.com
FAMILY : CPG
VERSION : 1.0
// Support: tech.team.motioncontrol@siemens.com
// Fax: +49 (0) 9131/98-1297
// stored: InstanceOfName EM01_00_Main
"EM01_00_Main"
BEGIN
END_DATA_BLOCK

// folder: EM02_Palletizing

DATA_BLOCK "EM02"   // DB31689
TITLE = EM02
{ S7_Optimized_Access := 'TRUE' }
AUTHOR : tech.team.motioncontrol@siemens.com
FAMILY : CPG
VERSION : 1.0
// Support: tech.team.motioncontrol@siemens.com
// Fax: +49 (0) 9131/98-1297
   VAR
      PackML_Sts : Struct   // PackML Module Status - EM and all control modules
         Unit : "CPG_typePackML_ModuleSts";   // PackML Module Status - EM - master status
         Alarm : "CPG_typePackML_ModuleSts";   // PackML Module Status - alarm status
         CM01 : "CPG_typePackML_ModuleSts";   // PackML Module Status - CM 01
         CM02 : "CPG_typePackML_ModuleSts";   // PackML Module Status - CM 02
         CM03 : "CPG_typePackML_ModuleSts";   // PackML Module Status - CM 03
         CM04 : "CPG_typePackML_ModuleSts";   // PackML Module Status - CM 04
         CM05 : "CPG_typePackML_ModuleSts";   // PackML Module Status - CM 05
         CM06 : "CPG_typePackML_ModuleSts";   // PackML Module Status - CM 06
         CM07 : "CPG_typePackML_ModuleSts";   // PackML Module Status - CM 07
         CM08 : "CPG_typePackML_ModuleSts";   // PackML Module Status - CM 08
         CM09 : "CPG_typePackML_ModuleSts";   // PackML Module Status - CM 09
         CM10 : "CPG_typePackML_ModuleSts";   // PackML Module Status - CM 10
      END_STRUCT;
      Alarm : "CPG_typeEventStatus";   // Alarm Event Status - EM02 Status
      Warning : "CPG_typeEventStatus";   // Warning Event Status - EM02 Status
      Status : "CPG_typeEventStatus";   // Event Status - EM02 Status
   END_VAR
BEGIN
END_DATA_BLOCK

// folder: EM02_Palletizing/Instances

DATA_BLOCK "InstEM02_00_Main"   // DB31680
TITLE = InstEM02_00_Main
{ S7_Optimized_Access := 'TRUE' }
AUTHOR : tech.team.motioncontrol@siemens.com
FAMILY : CPG
VERSION : 1.0
// Support: tech.team.motioncontrol@siemens.com
// Fax: +49 (0) 9131/98-1297
// stored: InstanceOfName EM02_00_Main
"EM02_00_Main"
BEGIN
END_DATA_BLOCK

// folder: GlobalData

DATA_BLOCK "Controls"   // DB1
{ S7_Optimized_Access := 'TRUE' }
VERSION : 0.1
   VAR
      Input : Bool;
      Reset : Bool;
      Timeout : Time;
      "Counter" : Int;
      NO_OF_LAYERS : Int;
   END_VAR
BEGIN
END_DATA_BLOCK

DATA_BLOCK "Alarm"   // DB31610
TITLE = CPG_Alarm
{ S7_Optimized_Access := 'TRUE' }
AUTHOR : tech.team.motioncontrol@siemens.com
FAMILY : CPG
VERSION : 1.0
// Support: tech.team.motioncontrol@siemens.com
// Fax: +49 (0) 9131/98-1297
   VAR
      Summation : "CPG_typeEventSummation";   // Unit Mode - Event Summation
   END_VAR
BEGIN
   Summation.wrk_EventArraySize := 30;
END_DATA_BLOCK

DATA_BLOCK "Warning"   // DB31611
TITLE = CPG_Warning
{ S7_Optimized_Access := 'TRUE' }
AUTHOR : tech.team.motioncontrol@siemens.com
FAMILY : CPG
VERSION : 1.0
// Support: tech.team.motioncontrol@siemens.com
// Fax: +49 (0) 9131/98-1297
   VAR
      Summation : "CPG_typeEventSummation";   // Unit Mode - Warning Summation
   END_VAR
BEGIN
   Summation.wrk_EventArraySize := 30;
END_DATA_BLOCK

DATA_BLOCK "Status"   // DB31612
TITLE = CPG_Status
{ S7_Optimized_Access := 'TRUE' }
AUTHOR : tech.team.motioncontrol@siemens.com
FAMILY : CPG